(* Logix 5000 project; controller PLC_MCC1300_75F1 vendor 1 type 14 code 166 rev 32.11; software revision 32.04; part 36 of 83 *)
(* tags used below, declared in another part *)
   N12 : DINT[500];
   N16 : DINT[500];
   N17 : DINT[100];
   N601 : DINT[25];
   N602 : DINT[25];
   N603 : DINT[25];
   N604 : DINT[25];
   N605 : DINT[25];
   N606 : DINT[25];
   N607 : DINT[25];
   N608 : DINT[25];
   N609 : DINT[25];
   N610 : DINT[25];
   N611 : DINT[25];
   N612 : DINT[25];
   N613 : DINT[25];
   N614 : DINT[25];
   N615 : DINT[25];
   N616 : DINT[25];
   N617 : DINT[25];
   N618 : DINT[25];
   N619 : DINT[25];
   N620 : DINT[25];
   N621 : DINT[25];
   N622 : DINT[25];
   N623 : DINT[25];
   N624 : DINT[25];
   N625 : DINT[25];
   N626 : DINT[25];
   N627 : DINT[25];
   N628 : DINT[25];
   N629 : DINT[25];
   N630 : DINT[25];
   N631 : DINT[25];
   N632 : DINT[25];
   N633 : DINT[25];
   N634 : DINT[25];
   N635 : DINT[25];
   N636 : DINT[25];
   N637 : DINT[25];
   N638 : DINT[25];
   N639 : DINT[25];
   N640 : DINT[25];
   N641 : DINT[25];
   N642 : DINT[25];
   N643 : DINT[25];
   N644 : DINT[25];
   N645 : DINT[25];
   N646 : DINT[25];
   N647 : DINT[25];
   N648 : DINT[25];
   N649 : DINT[25];
   N650 : DINT[25];
   N651 : DINT[25];
   N652 : DINT[25];
   N653 : DINT[25];
   N654 : DINT[25];
   N655 : DINT[25];
   N656 : DINT[25];
   N657 : DINT[25];
   N658 : DINT[25];
   N659 : DINT[25];
   N660 : DINT[25];
   N662 : DINT[25];
   N663 : DINT[25];
   N664 : DINT[25];
   N665 : DINT[25];
   N666 : DINT[25];
   N667 : DINT[25];
   N668 : DINT[25];
   N669 : DINT[25];
   N670 : DINT[25];
   N671 : DINT[25];
   N672 : DINT[25];
   N673 : DINT[25];
   N674 : DINT[25];
   N675 : DINT[25];
   N676 : DINT[25];
   N677 : DINT[25];
   N678 : DINT[25];
   N679 : DINT[25];
   N680 : DINT[25];
   N681 : DINT[25];
   N682 : DINT[25];
   N683 : DINT[25];
   N684 : DINT[25];
   N685 : DINT[25];
   N686 : DINT[25];
   N687 : DINT[25];
   N688 : DINT[25];
   N689 : DINT[25];
   N690 : DINT[25];
   N691 : DINT[25];
   N692 : DINT[25];
   N693 : DINT[25];
   N694 : DINT[25];
   N695 : DINT[25];
   N696 : DINT[25];
   N697 : DINT[25];
   N698 : DINT[25];
   N699 : DINT[25];
   N7 : DINT[101];
   N700 : DINT[25];
   N701 : DINT[25];
   N702 : DINT[25];
   N703 : DINT[25];
   N704 : DINT[25];
   N705 : DINT[25];
   N706 : DINT[25];
   N707 : DINT[25];
   N708 : DINT[25];
   N709 : DINT[25];
   N710 : DINT[25];
   N711 : DINT[25];
   N712 : DINT[25];
   N713 : DINT[25];
   N714 : DINT[25];
   N715 : DINT[25];
   N716 : DINT[25];
   N717 : DINT[25];
   N718 : DINT[25];
   N719 : DINT[25];
   N720 : DINT[25];
   N721 : DINT[25];
   N723 : DINT[25];
   N724 : DINT[25];
   N725 : DINT[25];
   N726 : DINT[25];
   N727 : DINT[25];
   N728 : DINT[25];
   N729 : DINT[25];
   N730 : DINT[25];
   N731 : DINT[25];
   N732 : DINT[25];
   N733 : DINT[25];
   N734 : DINT[25];
   N735 : DINT[25];
   N736 : DINT[25];
   N737 : DINT[25];
   N738 : DINT[25];
   N739 : DINT[25];
   N740 : DINT[25];
   N741 : DINT[25];
   N742 : DINT[25];
   N743 : DINT[25];
   N744 : DINT[25];
   N745 : DINT[25];
   N746 : DINT[25];
   N747 : DINT[25];
   N748 : DINT[25];
   N749 : DINT[25];
   N750 : DINT[25];
   N751 : DINT[25];
   N752 : DINT[25];
   N753 : DINT[25];
   N754 : DINT[25];
   N755 : DINT[25];
   N756 : DINT[25];
   N758 : DINT[25];
   N759 : DINT[25];
   N760 : DINT[25];
   N761 : DINT[25];
   N762 : DINT[25];
   N763 : DINT[25];
   N764 : DINT[25];
   N765 : DINT[25];
   N766 : DINT[25];
   N767 : DINT[25];
   N768 : DINT[25];
   N769 : DINT[25];
   N770 : DINT[25];
   N771 : DINT[25];
   N772 : DINT[25];
   N773 : DINT[25];
   N774 : DINT[25];
   N775 : DINT[25];
   N776 : DINT[25];
   N777 : DINT[25];
   N778 : DINT[25];
   N779 : DINT[25];
   N780 : DINT[25];
   N781 : DINT[25];
   N782 : DINT[25];
   N783 : DINT[25];
   N784 : DINT[25];
   N785 : DINT[25];
   N786 : DINT[25];
   N787 : DINT[25];
   N788 : DINT[25];
   N789 : DINT[25];
   N790 : DINT[25];
   N791 : DINT[25];
   N792 : DINT[25];
   N793 : DINT[25];
   N794 : DINT[25];
   N795 : DINT[25];
   N796 : DINT[25];
   N797 : DINT[25];
   N798 : DINT[25];
   N799 : DINT[25];
   TMP_dDestFile : DINT;
   TMP_dDestOffset : DINT;
   TMP_dErrDestFile : DINT;
   TMP_dErrSourceFile : DINT;
   TMP_dNumValues : DINT;
   TMP_dSourceFile : DINT;
   TMP_dSourceOffset : DINT;
(* MainProgram, continued *)

ROUTINE _942_SbrCOP_ValFromFile   (* structured text *)
// This Task replaces [COP] functions containing expressions with data pointing. It is necessary to correctly parameterize the INPUT_Par which the function will then copy the values written in the parameters for the preset Length number depending on the case.
// V1.1
   
   SBR(TMP_dSourceFile, TMP_dSourceOffset, TMP_dDestFile, TMP_dDestOffset, TMP_dNumValues);
   
   TMP_dErrSourceFile := 0;
   TMP_dErrDestFile := 0;
   
   (*
   ////CAPIDINDEX N7
   	IF (TMP_dSourceFile = 7) AND (TMP_dDestFile = 601) THEN
   		COP(N7[TMP_dSourceOffset], N601[TMP_dDestOffset], TMP_dNumValues);
   	ELSIF (TMP_dSourceFile = 7) AND (TMP_dDestFile = 602) THEN
   		COP(N7[TMP_dSourceOffset], N602[TMP_dDestOffset], TMP_dNumValues);
   	ELSIF (TMP_dSourceFile = 7) AND (TMP_dDestFile = 603) THEN
   		COP(N7[TMP_dSourceOffset], N603[TMP_dDestOffset], TMP_dNumValues);
   	ELSIF (TMP_dSourceFile = 7) AND (TMP_dDestFile = 604) THEN
   		COP(N7[TMP_dSourceOffset], N604[TMP_dDestOffset], TMP_dNumValues);
   	ELSIF (TMP_dSourceFile = 7) AND (TMP_dDestFile = 605) THEN
   		COP(N7[TMP_dSourceOffset], N605[TMP_dDestOffset], TMP_dNumValues);
   	ELSIF (TMP_dSourceFile = 7) AND (TMP_dDestFile = 606) THEN
   		COP(N7[TMP_dSourceOffset], N606[TMP_dDestOffset], TMP_dNumValues);
   	ELSIF (TMP_dSourceFile = 7) AND (TMP_dDestFile = 607) THEN
   		COP(N7[TMP_dSourceOffset], N607[TMP_dDestOffset], TMP_dNumValues);
   	ELSIF (TMP_dSourceFile = 7) AND (TMP_dDestFile = 608) THEN
   		COP(N7[TMP_dSourceOffset], N608[TMP_dDestOffset], TMP_dNumValues);
   	ELSIF (TMP_dSourceFile = 7) AND (TMP_dDestFile = 609) THEN
   		COP(N7[TMP_dSourceOffset], N609[TMP_dDestOffset], TMP_dNumValues);
   	ELSIF (TMP_dSourceFile = 7) AND (TMP_dDestFile = 610) THEN
   		COP(N7[TMP_dSourceOffset], N610[TMP_dDestOffset], TMP_dNumValues);
   	ELSIF (TMP_dSourceFile = 7) AND (TMP_dDestFile = 611) THEN
   		COP(N7[TMP_dSourceOffset], N611[TMP_dDestOffset], TMP_dNumValues);
   	ELSIF (TMP_dSourceFile = 7) AND (TMP_dDestFile = 612) THEN
   		COP(N7[TMP_dSourceOffset], N612[TMP_dDestOffset], TMP_dNumValues);
   	ELSIF (TMP_dSourceFile = 7) AND (TMP_dDestFile = 613) THEN
   		COP(N7[TMP_dSourceOffset], N613[TMP_dDestOffset], TMP_dNumValues);
   	ELSIF (TMP_dSourceFile = 7) AND (TMP_dDestFile = 614) THEN
   		COP(N7[TMP_dSourceOffset], N614[TMP_dDestOffset], TMP_dNumValues);
   	ELSIF (TMP_dSourceFile = 7) AND (TMP_dDestFile = 615) THEN
   		COP(N7[TMP_dSourceOffset], N615[TMP_dDestOffset], TMP_dNumValues);
   	ELSIF (TMP_dSourceFile = 7) AND (TMP_dDestFile = 616) THEN
   		COP(N7[TMP_dSourceOffset], N616[TMP_dDestOffset], TMP_dNumValues);
   	ELSIF (TMP_dSourceFile = 7) AND (TMP_dDestFile = 617) THEN
   		COP(N7[TMP_dSourceOffset], N617[TMP_dDestOffset], TMP_dNumValues);
   	ELSIF (TMP_dSourceFile = 7) AND (TMP_dDestFile = 618) THEN
   		COP(N7[TMP_dSourceOffset], N618[TMP_dDestOffset], TMP_dNumValues);
   	ELSIF (TMP_dSourceFile = 7) AND (TMP_dDestFile = 619) THEN
   		COP(N7[TMP_dSourceOffset], N619[TMP_dDestOffset], TMP_dNumValues);
   	ELSIF (TMP_dSourceFile = 7) AND (TMP_dDestFile = 620) THEN
   		COP(N7[TMP_dSourceOffset], N620[TMP_dDestOffset], TMP_dNumValues);
   	ELSIF (TMP_dSourceFile = 7) AND (TMP_dDestFile = 621) THEN
   		COP(N7[TMP_dSourceOffset], N621[TMP_dDestOffset], TMP_dNumValues);
   	ELSIF (TMP_dSourceFile = 7) AND (TMP_dDestFile = 622) THEN
   		COP(N7[TMP_dSourceOffset], N622[TMP_dDestOffset], TMP_dNumValues);
   	ELSIF (TMP_dSourceFile = 7) AND (TMP_dDestFile = 623) THEN
   		COP(N7[TMP_dSourceOffset], N623[TMP_dDestOffset], TMP_dNumValues);
   	ELSIF (TMP_dSourceFile = 7) AND (TMP_dDestFile = 624) THEN
   		COP(N7[TMP_dSourceOffset], N624[TMP_dDestOffset], TMP_dNumValues);
   	ELSIF (TMP_dSourceFile = 7) AND (TMP_dDestFile = 625) THEN
   		COP(N7[TMP_dSourceOffset], N625[TMP_dDestOffset], TMP_dNumValues);
   	ELSIF (TMP_dSourceFile = 7) AND (TMP_dDestFile = 626) THEN
   		COP(N7[TMP_dSourceOffset], N626[TMP_dDestOffset], TMP_dNumValues);
   	ELSIF (TMP_dSourceFile = 7) AND (TMP_dDestFile = 627) THEN
   		COP(N7[TMP_dSourceOffset], N627[TMP_dDestOffset], TMP_dNumValues);
   	ELSIF (TMP_dSourceFile = 7) AND (TMP_dDestFile = 628) THEN
   		COP(N7[TMP_dSourceOffset], N628[TMP_dDestOffset], TMP_dNumValues);
   	ELSIF (TMP_dSourceFile = 7) AND (TMP_dDestFile = 629) THEN
   		COP(N7[TMP_dSourceOffset], N629[TMP_dDestOffset], TMP_dNumValues);
   	ELSIF (TMP_dSourceFile = 7) AND (TMP_dDestFile = 630) THEN
   		COP(N7[TMP_dSourceOffset], N630[TMP_dDestOffset], TMP_dNumValues);
   	ELSIF (TMP_dSourceFile = 7) AND (TMP_dDestFile = 631) THEN
   		COP(N7[TMP_dSourceOffset], N631[TMP_dDestOffset], TMP_dNumValues);
   	ELSIF (TMP_dSourceFile = 7) AND (TMP_dDestFile = 632) THEN
   		COP(N7[TMP_dSourceOffset], N632[TMP_dDestOffset], TMP_dNumValues);
   	ELSIF (TMP_dSourceFile = 7) AND (TMP_dDestFile = 633) THEN
   		COP(N7[TMP_dSourceOffset], N633[TMP_dDestOffset], TMP_dNumValues);
   	ELSIF (TMP_dSourceFile = 7) AND (TMP_dDestFile = 634) THEN
   		COP(N7[TMP_dSourceOffset], N634[TMP_dDestOffset], TMP_dNumValues);
   	ELSIF (TMP_dSourceFile = 7) AND (TMP_dDestFile = 635) THEN
   		COP(N7[TMP_dSourceOffset], N635[TMP_dDestOffset], TMP_dNumValues);
   	ELSIF (TMP_dSourceFile = 7) AND (TMP_dDestFile = 636) THEN
   		COP(N7[TMP_dSourceOffset], N636[TMP_dDestOffset], TMP_dNumValues);
   	ELSIF (TMP_dSourceFile = 7) AND (TMP_dDestFile = 637) THEN
   		COP(N7[TMP_dSourceOffset], N637[TMP_dDestOffset], TMP_dNumValues);
   	ELSIF (TMP_dSourceFile = 7) AND (TMP_dDestFile = 638) THEN
   		COP(N7[TMP_dSourceOffset], N638[TMP_dDestOffset], TMP_dNumValues);
   	ELSIF (TMP_dSourceFile = 7) AND (TMP_dDestFile = 639) THEN
   		COP(N7[TMP_dSourceOffset], N639[TMP_dDestOffset], TMP_dNumValues);
   	ELSIF (TMP_dSourceFile = 7) AND (TMP_dDestFile = 640) THEN
   		COP(N7[TMP_dSourceOffset], N640[TMP_dDestOffset], TMP_dNumValues);
   	ELSIF (TMP_dSourceFile = 7) AND (TMP_dDestFile = 641) THEN
   		COP(N7[TMP_dSourceOffset], N641[TMP_dDestOffset], TMP_dNumValues);
   	ELSIF (TMP_dSourceFile = 7) AND (TMP_dDestFile = 642) THEN
   		COP(N7[TMP_dSourceOffset], N642[TMP_dDestOffset], TMP_dNumValues);
   	ELSIF (TMP_dSourceFile = 7) AND (TMP_dDestFile = 643) THEN
   		COP(N7[TMP_dSourceOffset], N643[TMP_dDestOffset], TMP_dNumValues);
   	ELSIF (TMP_dSourceFile = 7) AND (TMP_dDestFile = 644) THEN
   		COP(N7[TMP_dSourceOffset], N644[TMP_dDestOffset], TMP_dNumValues);
   	ELSIF (TMP_dSourceFile = 7) AND (TMP_dDestFile = 645) THEN
   		COP(N7[TMP_dSourceOffset], N645[TMP_dDestOffset], TMP_dNumValues);
   	ELSIF (TMP_dSourceFile = 7) AND (TMP_dDestFile = 646) THEN
   		COP(N7[TMP_dSourceOffset], N646[TMP_dDestOffset], TMP_dNumValues);
   	ELSIF (TMP_dSourceFile = 7) AND (TMP_dDestFile = 647) THEN
   		COP(N7[TMP_dSourceOffset], N647[TMP_dDestOffset], TMP_dNumValues);
   	ELSIF (TMP_dSourceFile = 7) AND (TMP_dDestFile = 648) THEN
   		COP(N7[TMP_dSourceOffset], N648[TMP_dDestOffset], TMP_dNumValues);
   	ELSIF (TMP_dSourceFile = 7) AND (TMP_dDestFile = 649) THEN
   		COP(N7[TMP_dSourceOffset], N649[TMP_dDestOffset], TMP_dNumValues);
   	ELSIF (TMP_dSourceFile = 7) AND (TMP_dDestFile = 650) THEN
   		COP(N7[TMP_dSourceOffset], N650[TMP_dDestOffset], TMP_dNumValues);
   	ELSIF (TMP_dSourceFile = 7) AND (TMP_dDestFile = 651) THEN
   		COP(N7[TMP_dSourceOffset], N651[TMP_dDestOffset], TMP_dNumValues);
   	ELSIF (TMP_dSourceFile = 7) AND (TMP_dDestFile = 652) THEN
   		COP(N7[TMP_dSourceOffset], N652[TMP_dDestOffset], TMP_dNumValues);
   	ELSIF (TMP_dSourceFile = 7) AND (TMP_dDestFile = 653) THEN
   		COP(N7[TMP_dSourceOffset], N653[TMP_dDestOffset], TMP_dNumValues);
   	ELSIF (TMP_dSourceFile = 7) AND (TMP_dDestFile = 654) THEN
   		COP(N7[TMP_dSourceOffset], N654[TMP_dDestOffset], TMP_dNumValues);
   	ELSIF (TMP_dSourceFile = 7) AND (TMP_dDestFile = 655) THEN
   		COP(N7[TMP_dSourceOffset], N655[TMP_dDestOffset], TMP_dNumValues);
   	ELSIF (TMP_dSourceFile = 7) AND (TMP_dDestFile = 656) THEN
   		COP(N7[TMP_dSourceOffset], N656[TMP_dDestOffset], TMP_dNumValues);
   	ELSIF (TMP_dSourceFile = 7) AND (TMP_dDestFile = 657) THEN
   		COP(N7[TMP_dSourceOffset], N657[TMP_dDestOffset], TMP_dNumValues);
   	ELSIF (TMP_dSourceFile = 7) AND (TMP_dDestFile = 658) THEN
   		COP(N7[TMP_dSourceOffset], N658[TMP_dDestOffset], TMP_dNumValues);
   	ELSIF (TMP_dSourceFile = 7) AND (TMP_dDestFile = 659) THEN
   		COP(N7[TMP_dSourceOffset], N659[TMP_dDestOffset], TMP_dNumValues);
   	ELSIF (TMP_dSourceFile = 7) AND (TMP_dDestFile = 660) THEN
   		COP(N7[TMP_dSourceOffset], N660[TMP_dDestOffset], TMP_dNumValues);
   	ELSIF (TMP_dSourceFile = 7) AND (TMP_dDestFile = 661) THEN
   		COP(N7[TMP_dSourceOffset], N661[TMP_dDestOffset], TMP_dNumValues);
   	ELSIF (TMP_dSourceFile = 7) AND (TMP_dDestFile = 662) THEN
   		COP(N7[TMP_dSourceOffset], N662[TMP_dDestOffset], TMP_dNumValues);
   	ELSIF (TMP_dSourceFile = 7) AND (TMP_dDestFile = 663) THEN
   		COP(N7[TMP_dSourceOffset], N663[TMP_dDestOffset], TMP_dNumValues);
   	ELSIF (TMP_dSourceFile = 7) AND (TMP_dDestFile = 664) THEN
   		COP(N7[TMP_dSourceOffset], N664[TMP_dDestOffset], TMP_dNumValues);
   	ELSIF (TMP_dSourceFile = 7) AND (TMP_dDestFile = 665) THEN
   		COP(N7[TMP_dSourceOffset], N665[TMP_dDestOffset], TMP_dNumValues);
   	ELSIF (TMP_dSourceFile = 7) AND (TMP_dDestFile = 666) THEN
   		COP(N7[TMP_dSourceOffset], N666[TMP_dDestOffset], TMP_dNumValues);
   	ELSIF (TMP_dSourceFile = 7) AND (TMP_dDestFile = 667) THEN
   		COP(N7[TMP_dSourceOffset], N667[TMP_dDestOffset], TMP_dNumValues);
   	ELSIF (TMP_dSourceFile = 7) AND (TMP_dDestFile = 668) THEN
   		COP(N7[TMP_dSourceOffset], N668[TMP_dDestOffset], TMP_dNumValues);
   	ELSIF (TMP_dSourceFile = 7) AND (TMP_dDestFile = 669) THEN
   		COP(N7[TMP_dSourceOffset], N669[TMP_dDestOffset], TMP_dNumValues);
   	ELSIF (TMP_dSourceFile = 7) AND (TMP_dDestFile = 670) THEN
   		COP(N7[TMP_dSourceOffset], N670[TMP_dDestOffset], TMP_dNumValues);
   	ELSIF (TMP_dSourceFile = 7) AND (TMP_dDestFile = 671) THEN
   		COP(N7[TMP_dSourceOffset], N671[TMP_dDestOffset], TMP_dNumValues);
   	ELSIF (TMP_dSourceFile = 7) AND (TMP_dDestFile = 672) THEN
   		COP(N7[TMP_dSourceOffset], N672[TMP_dDestOffset], TMP_dNumValues);
   	ELSIF (TMP_dSourceFile = 7) AND (TMP_dDestFile = 673) THEN
   		COP(N7[TMP_dSourceOffset], N673[TMP_dDestOffset], TMP_dNumValues);
   	ELSIF (TMP_dSourceFile = 7) AND (TMP_dDestFile = 674) THEN
   		COP(N7[TMP_dSourceOffset], N674[TMP_dDestOffset], TMP_dNumValues);
   	ELSIF (TMP_dSourceFile = 7) AND (TMP_dDestFile = 675) THEN
   		COP(N7[TMP_dSourceOffset], N675[TMP_dDestOffset], TMP_dNumValues);
   	ELSIF (TMP_dSourceFile = 7) AND (TMP_dDestFile = 676) THEN
   		COP(N7[TMP_dSourceOffset], N676[TMP_dDestOffset], TMP_dNumValues);
   	ELSIF (TMP_dSourceFile = 7) AND (TMP_dDestFile = 677) THEN
   		COP(N7[TMP_dSourceOffset], N677[TMP_dDestOffset], TMP_dNumValues);
   	ELSIF (TMP_dSourceFile = 7) AND (TMP_dDestFile = 678) THEN
   		COP(N7[TMP_dSourceOffset], N678[TMP_dDestOffset], TMP_dNumValues);
   	ELSIF (TMP_dSourceFile = 7) AND (TMP_dDestFile = 679) THEN
   		COP(N7[TMP_dSourceOffset], N679[TMP_dDestOffset], TMP_dNumValues);
   	ELSIF (TMP_dSourceFile = 7) AND (TMP_dDestFile = 680) THEN
   		COP(N7[TMP_dSourceOffset], N680[TMP_dDestOffset], TMP_dNumValues);
   	ELSIF (TMP_dSourceFile = 7) AND (TMP_dDestFile = 681) THEN
   		COP(N7[TMP_dSourceOffset], N681[TMP_dDestOffset], TMP_dNumValues);
   	ELSIF (TMP_dSourceFile = 7) AND (TMP_dDestFile = 682) THEN
   		COP(N7[TMP_dSourceOffset], N682[TMP_dDestOffset], TMP_dNumValues);
   	ELSIF (TMP_dSourceFile = 7) AND (TMP_dDestFile = 683) THEN
   		COP(N7[TMP_dSourceOffset], N683[TMP_dDestOffset], TMP_dNumValues);
   	ELSIF (TMP_dSourceFile = 7) AND (TMP_dDestFile = 684) THEN
   		COP(N7[TMP_dSourceOffset], N684[TMP_dDestOffset], TMP_dNumValues);
   	ELSIF (TMP_dSourceFile = 7) AND (TMP_dDestFile = 685) THEN
   		COP(N7[TMP_dSourceOffset], N685[TMP_dDestOffset], TMP_dNumValues);
   	ELSIF (TMP_dSourceFile = 7) AND (TMP_dDestFile = 686) THEN
   		COP(N7[TMP_dSourceOffset], N686[TMP_dDestOffset], TMP_dNumValues);
   	ELSIF (TMP_dSourceFile = 7) AND (TMP_dDestFile = 687) THEN
   		COP(N7[TMP_dSourceOffset], N687[TMP_dDestOffset], TMP_dNumValues);
   	ELSIF (TMP_dSourceFile = 7) AND (TMP_dDestFile = 688) THEN
   		COP(N7[TMP_dSourceOffset], N688[TMP_dDestOffset], TMP_dNumValues);
   	ELSIF (TMP_dSourceFile = 7) AND (TMP_dDestFile = 689) THEN
   		COP(N7[TMP_dSourceOffset], N689[TMP_dDestOffset], TMP_dNumValues);
   	ELSIF (TMP_dSourceFile = 7) AND (TMP_dDestFile = 690) THEN
   		COP(N7[TMP_dSourceOffset], N690[TMP_dDestOffset], TMP_dNumValues);
   	ELSIF (TMP_dSourceFile = 7) AND (TMP_dDestFile = 691) THEN
   		COP(N7[TMP_dSourceOffset], N691[TMP_dDestOffset], TMP_dNumValues);
   	ELSIF (TMP_dSourceFile = 7) AND (TMP_dDestFile = 692) THEN
   		COP(N7[TMP_dSourceOffset], N692[TMP_dDestOffset], TMP_dNumValues);
   	ELSIF (TMP_dSourceFile = 7) AND (TMP_dDestFile = 693) THEN
   		COP(N7[TMP_dSourceOffset], N693[TMP_dDestOffset], TMP_dNumValues);
   	ELSIF (TMP_dSourceFile = 7) AND (TMP_dDestFile = 694) THEN
   		COP(N7[TMP_dSourceOffset], N694[TMP_dDestOffset], TMP_dNumValues);
   	ELSIF (TMP_dSourceFile = 7) AND (TMP_dDestFile = 695) THEN
   		COP(N7[TMP_dSourceOffset], N695[TMP_dDestOffset], TMP_dNumValues);
   	ELSIF (TMP_dSourceFile = 7) AND (TMP_dDestFile = 696) THEN
   		COP(N7[TMP_dSourceOffset], N696[TMP_dDestOffset], TMP_dNumValues);
   	ELSIF (TMP_dSourceFile = 7) AND (TMP_dDestFile = 697) THEN
   		COP(N7[TMP_dSourceOffset], N697[TMP_dDestOffset], TMP_dNumValues);
   	ELSIF (TMP_dSourceFile = 7) AND (TMP_dDestFile = 698) THEN
   		COP(N7[TMP_dSourceOffset], N698[TMP_dDestOffset], TMP_dNumValues);
   	ELSIF (TMP_dSourceFile = 7) AND (TMP_dDestFile = 699) THEN
   		COP(N7[TMP_dSourceOffset], N699[TMP_dDestOffset], TMP_dNumValues);
   	ELSIF (TMP_dSourceFile = 7) AND (TMP_dDestFile = 700) THEN
   		COP(N7[TMP_dSourceOffset], N700[TMP_dDestOffset], TMP_dNumValues);
   	ELSIF (TMP_dSourceFile = 7) AND (TMP_dDestFile = 701) THEN
   		COP(N7[TMP_dSourceOffset], N701[TMP_dDestOffset], TMP_dNumValues);
   	ELSIF (TMP_dSourceFile = 7) AND (TMP_dDestFile = 702) THEN
   		COP(N7[TMP_dSourceOffset], N702[TMP_dDestOffset], TMP_dNumValues);
   	ELSIF (TMP_dSourceFile = 7) AND (TMP_dDestFile = 703) THEN
   		COP(N7[TMP_dSourceOffset], N703[TMP_dDestOffset], TMP_dNumValues);
   	ELSIF (TMP_dSourceFile = 7) AND (TMP_dDestFile = 704) THEN
   		COP(N7[TMP_dSourceOffset], N704[TMP_dDestOffset], TMP_dNumValues);
   	ELSIF (TMP_dSourceFile = 7) AND (TMP_dDestFile = 705) THEN
   		COP(N7[TMP_dSourceOffset], N705[TMP_dDestOffset], TMP_dNumValues);
   	ELSIF (TMP_dSourceFile = 7) AND (TMP_dDestFile = 706) THEN
   		COP(N7[TMP_dSourceOffset], N706[TMP_dDestOffset], TMP_dNumValues);
   	ELSIF (TMP_dSourceFile = 7) AND (TMP_dDestFile = 707) THEN
   		COP(N7[TMP_dSourceOffset], N707[TMP_dDestOffset], TMP_dNumValues);
   	ELSIF (TMP_dSourceFile = 7) AND (TMP_dDestFile = 708) THEN
   		COP(N7[TMP_dSourceOffset], N708[TMP_dDestOffset], TMP_dNumValues);
   	ELSIF (TMP_dSourceFile = 7) AND (TMP_dDestFile = 709) THEN
   		COP(N7[TMP_dSourceOffset], N709[TMP_dDestOffset], TMP_dNumValues);
   	ELSIF (TMP_dSourceFile = 7) AND (TMP_dDestFile = 710) THEN
   		COP(N7[TMP_dSourceOffset], N710[TMP_dDestOffset], TMP_dNumValues);
   	ELSIF (TMP_dSourceFile = 7) AND (TMP_dDestFile = 711) THEN
   		COP(N7[TMP_dSourceOffset], N711[TMP_dDestOffset], TMP_dNumValues);
   	ELSIF (TMP_dSourceFile = 7) AND (TMP_dDestFile = 712) THEN
   		COP(N7[TMP_dSourceOffset], N712[TMP_dDestOffset], TMP_dNumValues);
   	ELSIF (TMP_dSourceFile = 7) AND (TMP_dDestFile = 713) THEN
   		COP(N7[TMP_dSourceOffset], N713[TMP_dDestOffset], TMP_dNumValues);
   	ELSIF (TMP_dSourceFile = 7) AND (TMP_dDestFile = 714) THEN
   		COP(N7[TMP_dSourceOffset], N714[TMP_dDestOffset], TMP_dNumValues);
   	ELSIF (TMP_dSourceFile = 7) AND (TMP_dDestFile = 715) THEN
   		COP(N7[TMP_dSourceOffset], N715[TMP_dDestOffset], TMP_dNumValues);
   	ELSIF (TMP_dSourceFile = 7) AND (TMP_dDestFile = 716) THEN
   		COP(N7[TMP_dSourceOffset], N716[TMP_dDestOffset], TMP_dNumValues);
   	ELSIF (TMP_dSourceFile = 7) AND (TMP_dDestFile = 717) THEN
   		COP(N7[TMP_dSourceOffset], N717[TMP_dDestOffset], TMP_dNumValues);
   	ELSIF (TMP_dSourceFile = 7) AND (TMP_dDestFile = 718) THEN
   		COP(N7[TMP_dSourceOffset], N718[TMP_dDestOffset], TMP_dNumValues);
   	ELSIF (TMP_dSourceFile = 7) AND (TMP_dDestFile = 719) THEN
   		COP(N7[TMP_dSourceOffset], N719[TMP_dDestOffset], TMP_dNumValues);
   	ELSIF (TMP_dSourceFile = 7) AND (TMP_dDestFile = 720) THEN
   		COP(N7[TMP_dSourceOffset], N720[TMP_dDestOffset], TMP_dNumValues);
   	ELSIF (TMP_dSourceFile = 7) AND (TMP_dDestFile = 721) THEN
   		COP(N7[TMP_dSourceOffset], N721[TMP_dDestOffset], TMP_dNumValues);
   	ELSIF (TMP_dSourceFile = 7) AND (TMP_dDestFile = 722) THEN
   		COP(N7[TMP_dSourceOffset], N722[TMP_dDestOffset], TMP_dNumValues);
   	ELSIF (TMP_dSourceFile = 7) AND (TMP_dDestFile = 723) THEN
   		COP(N7[TMP_dSourceOffset], N723[TMP_dDestOffset], TMP_dNumValues);
   	ELSIF (TMP_dSourceFile = 7) AND (TMP_dDestFile = 724) THEN
   		COP(N7[TMP_dSourceOffset], N724[TMP_dDestOffset], TMP_dNumValues);
   	ELSIF (TMP_dSourceFile = 7) AND (TMP_dDestFile = 725) THEN
   		COP(N7[TMP_dSourceOffset], N725[TMP_dDestOffset], TMP_dNumValues);
   	ELSIF (TMP_dSourceFile = 7) AND (TMP_dDestFile = 726) THEN
   		COP(N7[TMP_dSourceOffset], N726[TMP_dDestOffset], TMP_dNumValues);
   	ELSIF (TMP_dSourceFile = 7) AND (TMP_dDestFile = 727) THEN
   		COP(N7[TMP_dSourceOffset], N727[TMP_dDestOffset], TMP_dNumValues);
   	ELSIF (TMP_dSourceFile = 7) AND (TMP_dDestFile = 728) THEN
   		COP(N7[TMP_dSourceOffset], N728[TMP_dDestOffset], TMP_dNumValues);
   	ELSIF (TMP_dSourceFile = 7) AND (TMP_dDestFile = 729) THEN
   		COP(N7[TMP_dSourceOffset], N729[TMP_dDestOffset], TMP_dNumValues);
   	ELSIF (TMP_dSourceFile = 7) AND (TMP_dDestFile = 730) THEN
   		COP(N7[TMP_dSourceOffset], N730[TMP_dDestOffset], TMP_dNumValues);
   	ELSIF (TMP_dSourceFile = 7) AND (TMP_dDestFile = 731) THEN
   		COP(N7[TMP_dSourceOffset], N731[TMP_dDestOffset], TMP_dNumValues);
   	ELSIF (TMP_dSourceFile = 7) AND (TMP_dDestFile = 732) THEN
   		COP(N7[TMP_dSourceOffset], N732[TMP_dDestOffset], TMP_dNumValues);
   	ELSIF (TMP_dSourceFile = 7) AND (TMP_dDestFile = 733) THEN
   		COP(N7[TMP_dSourceOffset], N733[TMP_dDestOffset], TMP_dNumValues);
   	ELSIF (TMP_dSourceFile = 7) AND (TMP_dDestFile = 734) THEN
   		COP(N7[TMP_dSourceOffset], N734[TMP_dDestOffset], TMP_dNumValues);
   	ELSIF (TMP_dSourceFile = 7) AND (TMP_dDestFile = 735) THEN
   		COP(N7[TMP_dSourceOffset], N735[TMP_dDestOffset], TMP_dNumValues);
   	ELSIF (TMP_dSourceFile = 7) AND (TMP_dDestFile = 736) THEN
   		COP(N7[TMP_dSourceOffset], N736[TMP_dDestOffset], TMP_dNumValues);
   	ELSIF (TMP_dSourceFile = 7) AND (TMP_dDestFile = 737) THEN
   		COP(N7[TMP_dSourceOffset], N737[TMP_dDestOffset], TMP_dNumValues);
   	ELSIF (TMP_dSourceFile = 7) AND (TMP_dDestFile = 738) THEN
   		COP(N7[TMP_dSourceOffset], N738[TMP_dDestOffset], TMP_dNumValues);
   	ELSIF (TMP_dSourceFile = 7) AND (TMP_dDestFile = 739) THEN
   		COP(N7[TMP_dSourceOffset], N739[TMP_dDestOffset], TMP_dNumValues);
   	ELSIF (TMP_dSourceFile = 7) AND (TMP_dDestFile = 740) THEN
   		COP(N7[TMP_dSourceOffset], N740[TMP_dDestOffset], TMP_dNumValues);
   	ELSIF (TMP_dSourceFile = 7) AND (TMP_dDestFile = 741) THEN
   		COP(N7[TMP_dSourceOffset], N741[TMP_dDestOffset], TMP_dNumValues);
   	ELSIF (TMP_dSourceFile = 7) AND (TMP_dDestFile = 742) THEN
   		COP(N7[TMP_dSourceOffset], N742[TMP_dDestOffset], TMP_dNumValues);
   	ELSIF (TMP_dSourceFile = 7) AND (TMP_dDestFile = 743) THEN
   		COP(N7[TMP_dSourceOffset], N743[TMP_dDestOffset], TMP_dNumValues);
   	ELSIF (TMP_dSourceFile = 7) AND (TMP_dDestFile = 744) THEN
   		COP(N7[TMP_dSourceOffset], N744[TMP_dDestOffset], TMP_dNumValues);
   	ELSIF (TMP_dSourceFile = 7) AND (TMP_dDestFile = 745) THEN
   		COP(N7[TMP_dSourceOffset], N745[TMP_dDestOffset], TMP_dNumValues);
   	ELSIF (TMP_dSourceFile = 7) AND (TMP_dDestFile = 746) THEN
   		COP(N7[TMP_dSourceOffset], N746[TMP_dDestOffset], TMP_dNumValues);
   	ELSIF (TMP_dSourceFile = 7) AND (TMP_dDestFile = 747) THEN
   		COP(N7[TMP_dSourceOffset], N747[TMP_dDestOffset], TMP_dNumValues);
   	ELSIF (TMP_dSourceFile = 7) AND (TMP_dDestFile = 748) THEN
   		COP(N7[TMP_dSourceOffset], N748[TMP_dDestOffset], TMP_dNumValues);
   	ELSIF (TMP_dSourceFile = 7) AND (TMP_dDestFile = 749) THEN
   		COP(N7[TMP_dSourceOffset], N749[TMP_dDestOffset], TMP_dNumValues);
   	ELSIF (TMP_dSourceFile = 7) AND (TMP_dDestFile = 750) THEN
   		COP(N7[TMP_dSourceOffset], N750[TMP_dDestOffset], TMP_dNumValues);
   	ELSIF (TMP_dSourceFile = 7) AND (TMP_dDestFile = 751) THEN
   		COP(N7[TMP_dSourceOffset], N751[TMP_dDestOffset], TMP_dNumValues);
   	ELSIF (TMP_dSourceFile = 7) AND (TMP_dDestFile = 752) THEN
   		COP(N7[TMP_dSourceOffset], N752[TMP_dDestOffset], TMP_dNumValues);
   	ELSIF (TMP_dSourceFile = 7) AND (TMP_dDestFile = 753) THEN
   		COP(N7[TMP_dSourceOffset], N753[TMP_dDestOffset], TMP_dNumValues);
   	ELSIF (TMP_dSourceFile = 7) AND (TMP_dDestFile = 754) THEN
   		COP(N7[TMP_dSourceOffset], N754[TMP_dDestOffset], TMP_dNumValues);
   	ELSIF (TMP_dSourceFile = 7) AND (TMP_dDestFile = 755) THEN
   		COP(N7[TMP_dSourceOffset], N755[TMP_dDestOffset], TMP_dNumValues);
   	ELSIF (TMP_dSourceFile = 7) AND (TMP_dDestFile = 756) THEN
   		COP(N7[TMP_dSourceOffset], N756[TMP_dDestOffset], TMP_dNumValues);
   	ELSIF (TMP_dSourceFile = 7) AND (TMP_dDestFile = 757) THEN
   		COP(N7[TMP_dSourceOffset], N757[TMP_dDestOffset], TMP_dNumValues);
   	ELSIF (TMP_dSourceFile = 7) AND (TMP_dDestFile = 758) THEN
   		COP(N7[TMP_dSourceOffset], N758[TMP_dDestOffset], TMP_dNumValues);
   	ELSIF (TMP_dSourceFile = 7) AND (TMP_dDestFile = 759) THEN
   		COP(N7[TMP_dSourceOffset], N759[TMP_dDestOffset], TMP_dNumValues);
   	ELSIF (TMP_dSourceFile = 7) AND (TMP_dDestFile = 760) THEN
   		COP(N7[TMP_dSourceOffset], N760[TMP_dDestOffset], TMP_dNumValues);
   	ELSIF (TMP_dSourceFile = 7) AND (TMP_dDestFile = 761) THEN
   		COP(N7[TMP_dSourceOffset], N761[TMP_dDestOffset], TMP_dNumValues);
   	ELSIF (TMP_dSourceFile = 7) AND (TMP_dDestFile = 762) THEN
   		COP(N7[TMP_dSourceOffset], N762[TMP_dDestOffset], TMP_dNumValues);
   	ELSIF (TMP_dSourceFile = 7) AND (TMP_dDestFile = 763) THEN
   		COP(N7[TMP_dSourceOffset], N763[TMP_dDestOffset], TMP_dNumValues);
   	ELSIF (TMP_dSourceFile = 7) AND (TMP_dDestFile = 764) THEN
   		COP(N7[TMP_dSourceOffset], N764[TMP_dDestOffset], TMP_dNumValues);
   	ELSIF (TMP_dSourceFile = 7) AND (TMP_dDestFile = 765) THEN
   		COP(N7[TMP_dSourceOffset], N765[TMP_dDestOffset], TMP_dNumValues);
   	ELSIF (TMP_dSourceFile = 7) AND (TMP_dDestFile = 766) THEN
   		COP(N7[TMP_dSourceOffset], N766[TMP_dDestOffset], TMP_dNumValues);
   	ELSIF (TMP_dSourceFile = 7) AND (TMP_dDestFile = 767) THEN
   		COP(N7[TMP_dSourceOffset], N767[TMP_dDestOffset], TMP_dNumValues);
   	ELSIF (TMP_dSourceFile = 7) AND (TMP_dDestFile = 768) THEN
   		COP(N7[TMP_dSourceOffset], N768[TMP_dDestOffset], TMP_dNumValues);
   	ELSIF (TMP_dSourceFile = 7) AND (TMP_dDestFile = 769) THEN
   		COP(N7[TMP_dSourceOffset], N769[TMP_dDestOffset], TMP_dNumValues);
   	ELSIF (TMP_dSourceFile = 7) AND (TMP_dDestFile = 770) THEN
   		COP(N7[TMP_dSourceOffset], N770[TMP_dDestOffset], TMP_dNumValues);
   	ELSIF (TMP_dSourceFile = 7) AND (TMP_dDestFile = 771) THEN
   		COP(N7[TMP_dSourceOffset], N771[TMP_dDestOffset], TMP_dNumValues);
   	ELSIF (TMP_dSourceFile = 7) AND (TMP_dDestFile = 772) THEN
   		COP(N7[TMP_dSourceOffset], N772[TMP_dDestOffset], TMP_dNumValues);
   	ELSIF (TMP_dSourceFile = 7) AND (TMP_dDestFile = 773) THEN
   		COP(N7[TMP_dSourceOffset], N773[TMP_dDestOffset], TMP_dNumValues);
   	ELSIF (TMP_dSourceFile = 7) AND (TMP_dDestFile = 774) THEN
   		COP(N7[TMP_dSourceOffset], N774[TMP_dDestOffset], TMP_dNumValues);
   	ELSIF (TMP_dSourceFile = 7) AND (TMP_dDestFile = 775) THEN
   		COP(N7[TMP_dSourceOffset], N775[TMP_dDestOffset], TMP_dNumValues);
   	ELSIF (TMP_dSourceFile = 7) AND (TMP_dDestFile = 776) THEN
   		COP(N7[TMP_dSourceOffset], N776[TMP_dDestOffset], TMP_dNumValues);
   	ELSIF (TMP_dSourceFile = 7) AND (TMP_dDestFile = 777) THEN
   		COP(N7[TMP_dSourceOffset], N777[TMP_dDestOffset], TMP_dNumValues);
   	ELSIF (TMP_dSourceFile = 7) AND (TMP_dDestFile = 778) THEN
   		COP(N7[TMP_dSourceOffset], N778[TMP_dDestOffset], TMP_dNumValues);
   	ELSIF (TMP_dSourceFile = 7) AND (TMP_dDestFile = 779) THEN
   		COP(N7[TMP_dSourceOffset], N779[TMP_dDestOffset], TMP_dNumValues);
   	ELSIF (TMP_dSourceFile = 7) AND (TMP_dDestFile = 780) THEN
   		COP(N7[TMP_dSourceOffset], N780[TMP_dDestOffset], TMP_dNumValues);
   	ELSIF (TMP_dSourceFile = 7) AND (TMP_dDestFile = 781) THEN
   		COP(N7[TMP_dSourceOffset], N781[TMP_dDestOffset], TMP_dNumValues);
   	ELSIF (TMP_dSourceFile = 7) AND (TMP_dDestFile = 782) THEN
   		COP(N7[TMP_dSourceOffset], N782[TMP_dDestOffset], TMP_dNumValues);
   	ELSIF (TMP_dSourceFile = 7) AND (TMP_dDestFile = 783) THEN
   		COP(N7[TMP_dSourceOffset], N783[TMP_dDestOffset], TMP_dNumValues);
   	ELSIF (TMP_dSourceFile = 7) AND (TMP_dDestFile = 784) THEN
   		COP(N7[TMP_dSourceOffset], N784[TMP_dDestOffset], TMP_dNumValues);
   	ELSIF (TMP_dSourceFile = 7) AND (TMP_dDestFile = 785) THEN
   		COP(N7[TMP_dSourceOffset], N785[TMP_dDestOffset], TMP_dNumValues);
   	ELSIF (TMP_dSourceFile = 7) AND (TMP_dDestFile = 786) THEN
   		COP(N7[TMP_dSourceOffset], N786[TMP_dDestOffset], TMP_dNumValues);
   	ELSIF (TMP_dSourceFile = 7) AND (TMP_dDestFile = 787) THEN
   		COP(N7[TMP_dSourceOffset], N787[TMP_dDestOffset], TMP_dNumValues);
   	ELSIF (TMP_dSourceFile = 7) AND (TMP_dDestFile = 788) THEN
   		COP(N7[TMP_dSourceOffset], N788[TMP_dDestOffset], TMP_dNumValues);
   	ELSIF (TMP_dSourceFile = 7) AND (TMP_dDestFile = 789) THEN
   		COP(N7[TMP_dSourceOffset], N789[TMP_dDestOffset], TMP_dNumValues);
   	ELSIF (TMP_dSourceFile = 7) AND (TMP_dDestFile = 790) THEN
   		COP(N7[TMP_dSourceOffset], N790[TMP_dDestOffset], TMP_dNumValues);
   	ELSIF (TMP_dSourceFile = 7) AND (TMP_dDestFile = 791) THEN
   		COP(N7[TMP_dSourceOffset], N791[TMP_dDestOffset], TMP_dNumValues);
   	ELSIF (TMP_dSourceFile = 7) AND (TMP_dDestFile = 792) THEN
   		COP(N7[TMP_dSourceOffset], N792[TMP_dDestOffset], TMP_dNumValues);
   	ELSIF (TMP_dSourceFile = 7) AND (TMP_dDestFile = 793) THEN
   		COP(N7[TMP_dSourceOffset], N793[TMP_dDestOffset], TMP_dNumValues);
   	ELSIF (TMP_dSourceFile = 7) AND (TMP_dDestFile = 794) THEN
   		COP(N7[TMP_dSourceOffset], N794[TMP_dDestOffset], TMP_dNumValues);
   	ELSIF (TMP_dSourceFile = 7) AND (TMP_dDestFile = 795) THEN
   		COP(N7[TMP_dSourceOffset], N795[TMP_dDestOffset], TMP_dNumValues);
   	ELSIF (TMP_dSourceFile = 7) AND (TMP_dDestFile = 796) THEN
   		COP(N7[TMP_dSourceOffset], N796[TMP_dDestOffset], TMP_dNumValues);
   	ELSIF (TMP_dSourceFile = 7) AND (TMP_dDestFile = 797) THEN
   		COP(N7[TMP_dSourceOffset], N797[TMP_dDestOffset], TMP_dNumValues);
   	ELSIF (TMP_dSourceFile = 7) AND (TMP_dDestFile = 798) THEN
   		COP(N7[TMP_dSourceOffset], N798[TMP_dDestOffset], TMP_dNumValues);
   	ELSIF (TMP_dSourceFile = 7) AND (TMP_dDestFile = 799) THEN
   		COP(N7[TMP_dSourceOffset], N799[TMP_dDestOffset], TMP_dNumValues);